(* Logix 5000 project; controller MV vendor 1 type 14 code 217 rev 31.11; software revision 31.00; part 2 of 53 *)

   MC_N224 : INT[255] := ([0] := 70, [1] := 59, [2] := 96, [3] := -32768, [4] := 9999, [5] := 9999, [6] := 9999, [7] := -32768);   // P24 CHECK CIP program 24 plant item check list
   MC_N225 : INT[255] := ([0] := 70, [1] := 59, [2] := 96, [3] := -32768, [4] := 9999, [5] := 9999, [6] := 9999, [7] := -32768);   // P25 CHECK CIP program 25 plant item check list
   MC_N226 : INT[255] := ([0] := 79, [1] := -32768, [2] := 9999, [3] := 9999, [4] := 9999, [5] := 9999, [6] := 9999, [7] := -32768);   // P26 CHECK CIP program 26 plant item check list
   MC_N227 : INT[255] := ([0] := 62, [1] := 99, [2] := -32768, [3] := 9999, [4] := 9999, [5] := 9999, [6] := 9999, [7] := -32768);   // P27 CHECK CIP program 27 plant item check list
   MC_N228 : INT[255] := ([0] := 61, [1] := 98, [2] := -32768, [3] := 9999, [4] := 9999, [5] := 9999, [6] := 9999, [7] := -32768);   // P28 CHECK CIP program 28 plant item check list
   MC_N229 : INT[255] := ([0] := 60, [1] := 97, [2] := -32768, [3] := 9999, [4] := 9999, [5] := 9999, [6] := 9999, [7] := -32768);   // P29 CHECK CIP program 29 plant item check list
   MC_N23 : INT[255] := ([0] := -31733, [2] := 1500, [3] := 5, [7] := 5000, [11] := 100, [12] := 10, [13] := 20, [14] := 7, [15] := 1493, [17] := -819, [18] := 25828, [21] := 5042, [22] := 1500, [24] := 1500, [25] := 13106, [27] := 1500, [31] := 3, [34] := 23, [36] := 1493);   // P2 FLOW Control block and da ta for P2 flowrate P ID loop
        [37]   // P2 flowrate PID saved op.mode
        [31].1   // P2 flowrate PID loop high absolute alarm flag
        [14]   // P2 flowrate PID loop process variable
        [31].0   // P2 flowrate PID loop deviation alarm flag
        [28]   // P2 flowrate PID loop high absolute alarm setting
        [31].2   // P2 flowrate PID loop low absolute alarm flag
        [30]   // P2 flowrate PID loop deviation alarm setting
        [38]   // P2 flowrate PID saved PLC output
        [26]   // P2 flowrate PID loop PLC output
        [25]   // P2 flowrate PID loop local (PC) output
        [0].1   // P2 flowrate PID loop auto/manual flag
        [2]   // P2 flowrate PID loop setpoint
        [27]   // P2 flowrate PID loop PLC setpoint
        [29]   // P2 flowrate PID loop low absolute alarm setting
        [35]   // P2 flowrate PID loop desired output
        [23]   // P2 flow op.mode: 0: PLC manual; 1: PLC setpoint; 2: Local manual; 3: Local setpoint;
        [36]   // Work register
   MC_N230 : INT[255] := ([0] := 60, [1] := 97, [2] := -32768, [3] := 9999, [4] := 9999, [5] := 9999, [6] := 9999, [7] := -32768);   // P30 CHECK CIP program 30 plant item check list
   MC_N231 : INT[255] := ([0] := 60, [1] := 97, [2] := -32768, [3] := 9999, [4] := 9999, [5] := 9999, [6] := 9999, [7] := -32768);   // P31 CHECK CIP program 31 plant item check list
   MC_N232 : INT[255] := ([0] := 60, [1] := 97, [2] := -32768, [3] := 9999, [4] := 9999, [5] := 9999, [6] := 9999, [7] := -32768);   // P32 CHECK CIP program 32 plant item check list
   MC_N233 : INT[255] := ([0] := 59, [1] := 96, [2] := -32768, [3] := 9999, [4] := 9999, [5] := 9999, [6] := 9999, [7] := -32768);   // P33 CHECK CIP program 33 plant item check list
   MC_N234 : INT[255] := ([0] := 59, [1] := 96, [2] := -32768, [3] := 9999, [4] := 9999, [5] := 9999, [6] := 9999, [7] := -32768);   // P34 CHECK CIP program 34 plant item check list
   MC_N235 : INT[255] := ([0] := 59, [1] := 96, [2] := -32768, [3] := 9999, [4] := 9999, [5] := 9999, [6] := 9999, [7] := -32768);   // P35 CHECK CIP program 35 plant item check list
   MC_N236 : INT[255] := ([0] := 59, [1] := 96, [2] := -32768, [3] := 9999, [4] := 9999, [5] := 9999, [6] := 9999, [7] := -32768);   // P36 CHECK CIP program 36 plant item check list
   MC_N237 : INT[255] := ([0] := 59, [1] := 96, [2] := -32768, [3] := 9999, [4] := 9999, [5] := 9999, [6] := 9999, [7] := -32768);   // P37 CHECK CIP program 37 plant item check list
   MC_N238 : INT[255] := ([0] := 59, [1] := 96, [2] := -32768, [3] := 9999, [4] := 9999, [5] := 9999, [6] := 9999, [7] := -32768);   // P38 CHECK CIP program 38 plant item check list
   MC_N239 : INT[255] := ([0] := 59, [1] := 96, [2] := -32768, [3] := 9999, [4] := 9999, [5] := 9999, [6] := 9999, [7] := -32768);   // P39 CHECK CIP program 39 plant item check list
   MC_N245 : INT[255];   // CC_WORK Continuous checking program work area
        [4].11   // CW deenergised input flag
        [6]   // Checking timer accumulator mask
        [15].0   // Current checkword is unused flag
        [2]   // Current item's energised input pointer
        [1]   // Current item's output pointer
        [3]   // Current item's Deenergised input pointer
        [4].10   // CW energised input flag
        [10].0   // Checking scan enabled flag
        [4].9   // CW desired output flag
        [0]   // Checkword pointer
        [16]   // Output slot update counter
        [28]   // No.items checked this scan
        [4]   // Current item's checkword
        [4].13   // CW checking inhibit flag
        [27]   // No new faults counter
        [4].12   // CW cycle flag
        [4].15   // CW fault flag
        [4].8   // CW manual flag
   MC_N255 : INT[255] := ([0] := 2208, [1] := 2208, [2] := 2208, [3] := 2208, [4] := 2208, [5] := 1696, [6] := 2208, [7] := 2208, [8] := 2208, [9] := 2208, [10] := 2208, [11] := 1696, [12] := 2208, [13] := 2208, [14] := 1696, [15] := 2112, [16] := 1600, [17] := 2112, [18] := 2112, [19] := 10304, [20] := 2112, [21] := 2112, [22] := 2112, [23] := 2112, [24] := 2112, [25] := 10304, [26] := 2112, [27] := 2112, [28] := 2112, [29] := 2112, [30] := 2112, [31] := 2112, [32] := 2112, [33] := 2112, [34] := 2112, [35] := 2112, [36] := 2112, [37] := 2112, [38] := 2112, [39] := 2112, [40] := 2112, [41] := 2112, [42] := 2112, [43] := 2112, [44] := 2112, [45] := 2112, [46] := 2112, [47] := 2112, [48] := 2112, [49] := 2112, [50] := 2112, [51] := 2112, [52] := 8256, [53] := 8256, [55] := 8256, [56] := 2112, [59] := 2112, [60] := 2112, [61] := 2112, [62] := 2112,
        [63] := 2112, [64] := 1600, [65] := 2112, [66] := 1600, [67] := 2112, [68] := 2112, [69] := 2112, [70] := 2112, [71] := 2112, [72] := 2112, [73] := 2112, [74] := 2112, [75] := 2112, [76] := 2112, [77] := 2112, [78] := 2112, [79] := 2112, [96] := 1600, [97] := 1600, [98] := 1600, [99] := 1600);   // CHECKWORDS Plant item checkword s
   MC_N7 : INT[255] := ([0] := 23, [1] := 22, [2] := 28, [4] := 2005, [5] := 5, [6] := 563, [7] := 84, [8] := 657, [9] := 653, [10] := -1);   // INTEGER
        [6]   // CH1/PTX scaled input
        [7]   // CH2/PTX scaled input
        [2]   // CH1/CTX1 scaled input
        [3]   // CH2/CTX2 scaled input
        [0]   // DT1 CTX-001 scaled input
        [1]   // DT2 CTX-002 scaled input
        [8]   // DT1 TTX-001 scaled input
        [9]   // DT2 TTX-002 scaled input
        [10]   // CH2/FM FV Bypass scaled input
        [4]   // CH1/FM scaled input
        [5]   // CH2/FM scaled input
   MC_N80 : INT[255] := ([0] := 5, [1] := 50, [2] := 4, [6] := 3, [7] := 23, [8] := 650, [10] := -1, [11] := 1, [13] := 10800, [14] := 1, [17] := 50, [18] := 7, [19] := 1, [20] := 2, [21] := 18);   // SRV1_PLC Detergent tank 1 ser vice PLC data
        [13]   // SV1 event register
        [21].1   // Channel 1 DT1 in use flag
        [21].3   // Channel 2 DT1 in use flag
        [2].0   // DT1 service manual start button available
        [2].15   // DT1 service command update toggle flag
        [21].4   // CH1/DT1 maintain temp.during service flag
        [21].5   // CH2/DT1 maintain temp.during service flag
        [20]   // DT1 service command processor current step
        [2].4   // DT1 service abort button available
        [21].0   // CH1 request DT1 service flag
        [21].2   // CH2 request DT1 service flag
        [8]   // DT1 service target detergent temp.
        [2].1   // DT1 manual service startup in progress
        [18].8   // DT1 service drive caustic pump flag
        [18].0   // DT1 service active flag
        [32].0   // DT1 service start by boilerhouse OSR
        [2].3   // DT1 service continue button available
        [6].0   // DT1 detergent strength ok
        [10]   // DT1 service routine fault register
        [18].1   // DT1 automatic service flag
        [6].1   // DT1 detergent temperature ok
        [17]   // DT1 service restart step
        [18].2   // DT1 service complete
        [6].2   // DT1 detergent diluted
        [11]   // SV1 fault parameter #1
        [12]   // SV1 fault parameter #2
        [14]   // SV1 event parameter #1
        [15]   // SV1 event parameter #2
        [1]   // DT1 service current step
        [2].2   // DT1 service stop button available
        [7]   // DT1 service target detergent strength
        [18].14   // Reset DT1 service flag
        [0]   // DT1 Service status 0:Unavailable; 1:Idle; 2:Running; 3:Stopped; 4:Faulted 5: Automatic
   MC_N80_10_alarm : ALARM_DIGITAL;
   MC_N80_10_Alarm_Ready : BOOL;
   MC_N80_10_Delayed_Timer2 : TIMER := (PRE := 1000);
   MC_N80_10_Fault_Returned : STRING;
   MC_N80_10_SQL_Done : DINT := -1;
   MC_N80_13_alarm : ALARM_DIGITAL;
   MC_N80_13_Alarm_Ready : BOOL := 1;
   MC_N80_13_Delayed_Timer2 : TIMER := (PRE := 1000);
   MC_N80_13_Event_Returned : STRING := 'Detergent tank service complete.';
   MC_N80_13_SQL_Done : DINT := -1;
   MC_N80_19_0_Storagebit : BOOL;
   MC_N81 : INT[255];   // SV1_PC Detergent tank 1 ser vice PC to PLC data
        [0].2   // Stop DT1 service
        [0].15   // DT1 manual service startup cancelled
        [0].0   // DT1 initiate manual service startup
        [0].4   // Abort DT1 service
        [0].1   // Start DT1 manual service
        [0]   // DT1 service PC button selected
        [0].3   // Continue DT1 service
   MC_N82 : INT[255] := ([0] := 14, [1] := 16, [2] := 34, [3] := 36, [4] := 41, [5] := 43, [6] := 45, [7] := 66, [8] := 78, [9] := -32768, [10] := 9999, [11] := 9999, [12] := 9999, [13] := 9999, [14] := 9999, [15] := 9999);   // SV1 ITEMS Chwd.nos.of items to be checked for DT1 service
        [6]   // SV1 checkword no.
        [8]   // CP1 checkword no.
        [0]   // CH1/DR1 checkword no.
        [1]   // CH1/DT1 checkword no.
        [2]   // CH2/DR1 checkword no.
        [3]   // CH2/DT1 checkword no.
        [4]   // FL/D1 checkword no.
        [5]   // CD/T1 checkword no.
        [7]   // P3 checkword no.
   MC_N90 : INT[255] := ([0] := 1, [2] := -32767, [10] := -1, [11] := 2, [13] := 10800, [14] := 2);   // SV2_PLC Detergent tank 2 ser vice PLC data
        [13]   // SV2 event register
        [21].1   // Channel 1 DT2 in use flag
        [21].3   // Channel 2 DT2 in use flag
        [2].0   // DT2 service manual start button available
        [2].15   // DT2 service command update toggle flag
        [21].4   // CH1/DT2 maintain temp.during service flag
        [21].0   // CH1 request DT2 service flag
        [21].5   // CH2/DT2 maintain temp.during service flag
        [20]   // DT2 service command processor current step
        [21].2   // CH2 request DT2 service flag
        [8]   // DT2 service target detergent temp.
        [2].4   // DT2 service abort button available
        [18].0   // DT2 service active flag
        [2].1   // DT2 manual service startup in progress
        [32].0   // DT2 service start by boilerhouse OSR
        [18].8   // DT2 service drive caustic pump flag
        [2].3   // DT2 service continue button available
        [6].0   // DT2 detergent strength ok
        [10]   // DT2 service routine fault register
        [18].1   // DT2 automatic service flag
        [6].1   // DT2 detergent temperature ok
        [17]   // DT2 service restart step
        [18].2   // DT2 service complete
        [6].2   // DT2 detergent diluted
        [11]   // SV2 fault parameter #1
        [14]   // SV2 event parameter #1
        [1]   // DT2 service current step
        [2].2   // DT2 service stop button available
        [7]   // DT2 service target detergent strength
        [18].14   // Reset DT2 service flag
        [0]   // DT2 Service status 0:Unavailable; 1:Idle; 2:Running; 3:Stopped; 4:Faulted 5: Automatic
   MC_N90_10_alarm : ALARM_DIGITAL;
   MC_N90_10_Alarm_Ready : BOOL;
   MC_N90_10_Delayed_Timer2 : TIMER := (PRE := 1000);
   MC_N90_10_Fault_Returned : STRING;
   MC_N90_10_SQL_Done : DINT := -1;
   MC_N90_13_alarm : ALARM_DIGITAL;
   MC_N90_13_Alarm_Ready : BOOL := 1;
   MC_N90_13_Delayed_Timer2 : TIMER := (PRE := 1002);
   MC_N90_13_Event_Returned : STRING := 'Detergent tank service complete.';
   MC_N90_13_SQL_Done : DINT := -1;
   MC_N90_19_0_Storagebit : BOOL;
   MC_N90_32_0_Storagebit : BOOL;
   MC_N91 : INT[255];   // SV2_PC Detergent tank 2 ser vice PC to PLC data
        [0].2   // Stop DT2 service
        [0].15   // DT2 manual service startup cancelled
        [0].0   // DT2 initiate manual service startup
        [0].4   // Abort DT2 service
        [0].1   // Start DT2 manual service
        [0]   // DT2 service PC button selected
        [0].3   // Continue DT2 service
   MC_N92 : INT[255] := ([0] := 15, [1] := 17, [2] := 35, [3] := 37, [4] := 42, [5] := 44, [6] := 46, [7] := 67, [8] := 78, [9] := -32768, [10] := 9999, [11] := 9999, [12] := 9999, [13] := 9999, [14] := 9999, [15] := 9999);   // SV2 ITEMS Chwd.nos.of items to be checked for DT2 service
        [6]   // SV2 checkword no.
        [8]   // CP1 checkword no.
        [0]   // CH1/DR2 checkword no.
        [1]   // CH1/DT2 checkword no.
        [2]   // CH2/DR2 checkword no.
        [3]   // CH2/DT2 checkword no.
        [4]   // FL/D2 checkword no.
        [7]   // P4 checkword no.
        [5]   // CD/T2 checkword no.
   MC_ONE_SEC : ALIAS FOR MC_T4[0].DN;
   MC_P1 : PlantItem := (CW := 2#0000_0000_0000_0001_0000_1100_1000_1011, CheckTime := 8, CheckTimer := 8, DriveBits := 1);   // P1
   MC_P1_ALARM : ALARM_DIGITAL;
   MC_P1_D : ALIAS FOR RIO_Rack_2:10:O.Data.0;
   MC_P1_Flow_PID : PID := (CTL := -2139061120, EN := 1, PE := 1, INI := 1, DVNA := 1, PVHA := 1, SP := 200.0, KP := 0.5, KI := 50.0, MAXS := 500.0, SO := 72.11798, MAXO := 100.0, MINO := 10.0, UPD := 1.0, PV := 200.53125, ERR := -0.53125, OUT := 72.11798, MAXI := 500.0, TIE := 72.118, MAXCV := 100.0, MAXTIE := 100.0, DATA[0] := 72.171104, DATA[1] := -641.7, DATA[2] := 200.53125, DATA[3] := -0.53125, DATA[4] := 200.0, DATA[5] := 0.2, DATA[6] := 1.0, DATA[7] := 16.0, DATA[8] := 0.5, DATA[9] := 50.0, DATA[11] := 0.5, DATA[12] := 0.00016666666, DATA[15] := 1.0, DATA[16] := 1.0);
   MC_P1_Flow_PID_Output : REAL := 72.16245;
   MC_P1_FPID_RESTORE : ALIAS FOR MC_N100[29].4;
   MC_P1_FPID_SAVE : ALIAS FOR MC_N100[29].3;
   MC_P1_PPID_RESTORE : ALIAS FOR MC_N100[29].2;
   MC_P1_PPID_SAVE : ALIAS FOR MC_N100[29].1;
   MC_P1_Pressure_PID : PID := (CTL := -2071952768, EN := 1, SWM := 1, PE := 1, INI := 1, DVPA := 1, PVHA := 1, SP := 65.0, KP := 1.0, KI := 2.0, MAXS := 150.0, MAXO := 100.0, UPD := 1.0, PV := 52.26563, ERR := 12.734371, MAXI := 150.0, MAXCV := 100.0, MAXTIE := 100.0, DATA[0] := -8.489581, DATA[1] := -557.50006, DATA[2] := 52.26563, DATA[3] := 12.734371, DATA[4] := 65.0, DATA[5] := 0.6666667, DATA[6] := 1.0, DATA[7] := 16.0, DATA[8] := 1.0, DATA[9] := 2.0, DATA[11] := 1.0, DATA[12] := 0.008333334, DATA[15] := 1.0, DATA[16] := 1.0);
   MC_P1_Pressure_PID_Output : REAL;
   MC_P1_R : ALIAS FOR RIO_Rack_2:11:I.Data.0;
   MC_P1_SP_AO : PlantItem := (Scaled := 72.161766);   // P1_SP
   MC_P1_SP_AO_RawOutput : ALIAS FOR RIO_Rack_2:3:O.Ch0Data;   // Real Analog Input , Do Not Use In Code
   MC_P1_T : ALIAS FOR RIO_Rack_2:11:I.Data.15;
   MC_P2 : PlantItem := (CW := 2#0000_0000_0000_0000_0000_1100_0000_0000, CheckTime := 8, CheckTimer := 8);   // P2
   MC_P2_ALARM : ALARM_DIGITAL;
   MC_P2_D : ALIAS FOR RIO_Rack_2:10:O.Data.1;
   MC_P2_Flow_PID : PID := (CTL := -2071952768, EN := 1, SWM := 1, PE := 1, INI := 1, DVPA := 1, PVHA := 1, SP := 150.0, KP := 0.5, KI := 50.0, MAXS := 500.0, MAXO := 100.0, UPD := 1.0, PV := 1.0, ERR := 149.0, MAXI := 500.0, MAXCV := 100.0, MAXTIE := 100.0, DATA[0] := -14.900001, DATA[1] := -3.2, DATA[2] := 1.0, DATA[3] := 149.0, DATA[4] := 150.0, DATA[5] := 0.2, DATA[6] := 1.0, DATA[7] := 16.0, DATA[8] := 0.5, DATA[9] := 50.0, DATA[11] := 0.5, DATA[12] := 0.00016666666, DATA[15] := 1.0, DATA[16] := 1.0);
   MC_P2_Flow_PID_Output : REAL;
   MC_P2_FPID_RESTORE : ALIAS FOR MC_N120[29].4;
   MC_P2_FPID_SAVE : ALIAS FOR MC_N120[29].3;
   MC_P2_PPID_RESTORE : ALIAS FOR MC_N120[29].2;
   MC_P2_PPID_SAVE : ALIAS FOR MC_N120[29].1;
   MC_P2_Pressure_PID : PID := (CTL := -2071952768, EN := 1, SWM := 1, PE := 1, INI := 1, DVPA := 1, PVHA := 1, SP := 45.0, KP := 0.1, KI := 2.0, MAXS := 150.0, MAXO := 100.0, UPD := 1.0, PV := 8.3625, ERR := 36.6375, MAXI := 150.0, MAXCV := 100.0, MAXTIE := 100.0, DATA[0] := -2.4425, DATA[1] := -89.200005, DATA[2] := 8.3625, DATA[3] := 36.6375, DATA[4] := 45.0, DATA[5] := 0.6666667, DATA[6] := 1.0, DATA[7] := 16.0, DATA[8] := 0.1, DATA[9] := 2.0, DATA[11] := 0.1, DATA[12] := 0.00083333335, DATA[15] := 1.0, DATA[16] := 1.0);
   MC_P2_Pressure_PID_Output : REAL;
   MC_P2_R : ALIAS FOR RIO_Rack_2:11:I.Data.1;
   MC_P2_SP_AO : PlantItem;   // P2_SP
   MC_P2_SP_AO_RawOutput : ALIAS FOR RIO_Rack_2:3:O.Ch1Data;   // Real Analog Input , Do Not Use In Code
   MC_P2_T : ALIAS FOR RIO_Rack_2:11:I.Data.16;
   MC_P3 : PlantItem := (CW := 2#0000_0000_0000_0000_0000_1100_1000_1011, CheckTime := 8, CheckTimer := 8, DriveBits := 1);   // P3
   MC_P3_ALARM : ALARM_DIGITAL;
   MC_P3_D : ALIAS FOR RIO_Rack_2:10:O.Data.2;
   MC_P3_R : ALIAS FOR RIO_Rack_2:11:I.Data.2;
   MC_P4 : PlantItem := (CW := 2#0000_0000_0000_0000_0000_1100_0000_0000, CheckTime := 8, CheckTimer := 8);   // P4
   MC_P4_ALARM : ALARM_DIGITAL;
   MC_P4_D : ALIAS FOR RIO_Rack_2:10:O.Data.3;
   MC_P4_R : ALIAS FOR RIO_Rack_2:11:I.Data.3;
   MC_PILZ : PlantItem := (CW := 2#0000_0000_0000_0100_0000_0000_0000_0001);   // PILZ
   MC_PILZ_RawInput : ALIAS FOR RIO_Rack_2:12:I.Data.31;   // MC_PILZ
   MC_PROXY2 : PlantItem;   // PROXY2
   MC_PROXY2_RawInput : ALIAS FOR RIO_Rack_2:12:I.Data.30;   // MC_PROXY2
   MC_PROXY_RawInput : ALIAS FOR RIO_Rack_2:12:I.Data.14;   // MC_PROXY
   MC_PX_100 : PlantItem;   // PX_100
   MC_PX_100_RawInput : ALIAS FOR RIO_Rack_2:11:I.Data.18;   // MC_PX_100
   MC_PX_101 : PlantItem;   // PX_101
   MC_PX_101_RawInput : ALIAS FOR RIO_Rack_2:11:I.Data.19;   // MC_PX_101
   MC_R2_SW1 : PlantItem;   // R2_SW1
   MC_R2_SW1_RawInput : ALIAS FOR RIO_Rack_2:12:I.Data.0;   // MC_R2_SW1
   MC_R2_SW2 : PlantItem;   // R2_SW2
   MC_R2_SW2_RawInput : ALIAS FOR RIO_Rack_2:12:I.Data.1;   // MC_R2_SW2
   MC_R2_SW3 : PlantItem;   // R2_SW3
   MC_R2_SW3_1 : PlantItem;   // R2_SW3_1
   MC_R2_SW3_1_RawInput : ALIAS FOR RIO_Rack_2:12:I.Data.3;   // MC_R2_SW3_1
   MC_R2_SW3_RawInput : ALIAS FOR RIO_Rack_2:12:I.Data.2;   // MC_R2_SW3
   MC_R2_SW4 : PlantItem := (CW := 2#0000_0000_0000_0100_0000_0000_0000_0001);   // R2_SW4
   MC_R2_SW4_RawInput : ALIAS FOR RIO_Rack_2:12:I.Data.4;   // MC_R2_SW4
   MC_R3_SW1 : PlantItem;   // R3_SW1
   MC_R3_SW1_RawInput : ALIAS FOR RIO_Rack_2:12:I.Data.5;   // MC_R3_SW1
   MC_R3_SW2 : PlantItem;   // R3_SW2
   MC_R3_SW2_1 : PlantItem := (CW := 2#0000_0000_0000_0100_0000_0000_0010_0001);   // PROXY
   MC_R3_SW2_RawInput : ALIAS FOR RIO_Rack_2:12:I.Data.6;   // MC_R3_SW2
   MC_R3_SW3 : PlantItem;   // R3_SW3
   MC_R3_SW3_1 : ALIAS FOR MC_N112[9].1;
   MC_R3_SW3_2 : ALIAS FOR MC_N112[9].0;
   MC_R3_SW3_3 : ALIAS FOR MC_N112[9].2;
   MC_R3_SW3_RawInput : ALIAS FOR RIO_Rack_2:12:I.Data.7;   // MC_R3_SW3
   MC_R3R_C_ALARM : ALARM_DIGITAL;
   MC_R3R_DR : PlantItem := (CW := 2#0000_0000_0000_0000_0000_0000_0001_0000, CheckTime := 8, CheckTimer := 15);   // R3R_DR
   MC_R3R_DR_ALARM : ALARM_DIGITAL;
   MC_R3R_DR_C : ALIAS FOR RIO_Rack_2:9:I.Data.20;
   MC_R3R_DR_DR : ALIAS FOR RIO_Rack_2:8:O.Data.24;
   MC_R3R_DR_O : ALIAS FOR RIO_Rack_2:9:I.Data.16;
   MC_R3R_O_ALARM : ALARM_DIGITAL;
   MC_R3S_C_ALARM : ALARM_DIGITAL;
   MC_R3S_DR : PlantItem := (CW := 2#0000_0000_0000_0000_0000_0001_0000_0000, CheckTime := 8, CheckTimer := 15);   // R3S_DR
   MC_R3S_DR_ALARM : ALARM_DIGITAL;
   MC_R3S_DR_C : ALIAS FOR RIO_Rack_2:9:I.Data.15;
   MC_R3S_DR_DR : ALIAS FOR RIO_Rack_2:8:O.Data.23;
   MC_R3S_DR_O : ALIAS FOR RIO_Rack_2:9:I.Data.11;
   MC_R3S_O_ALARM : ALARM_DIGITAL;
   MC_R3V1 : PlantItem := (CW := 2#0000_0000_0000_0000_0000_0001_0000_0000, CheckTime := 8, CheckTimer := 15);   // R3V1
   MC_R3V1_ALARM : ALARM_DIGITAL;
   MC_R3V1_C : ALIAS FOR RIO_Rack_2:9:I.Data.12;
   MC_R3V1_DR : ALIAS FOR RIO_Rack_2:8:O.Data.20;
   MC_R3V1_O : ALIAS FOR RIO_Rack_2:9:I.Data.8;
   MC_R3V2 : PlantItem := (CW := 2#0000_0000_0000_0000_0000_0001_0000_0000, CheckTime := 8, CheckTimer := 15);   // R3V2
   MC_R3V2_ALARM : ALARM_DIGITAL;
   MC_R3V2_C : ALIAS FOR RIO_Rack_2:9:I.Data.13;
   MC_R3V2_DR : ALIAS FOR RIO_Rack_2:8:O.Data.21;
   MC_R3V2_O : ALIAS FOR RIO_Rack_2:9:I.Data.9;
   MC_R3V3_C : ALIAS FOR RIO_Rack_2:9:I.Data.14;
   MC_R3V3_O : ALIAS FOR RIO_Rack_2:9:I.Data.10;
   MC_R4_SW1 : PlantItem;   // R4_SW1
   MC_R4_SW1_RawInput : ALIAS FOR RIO_Rack_2:12:I.Data.8;   // MC_R4_SW1
   MC_R4_SW2 : PlantItem;   // R4_SW2
   MC_R4_SW2_RawInput : ALIAS FOR RIO_Rack_2:12:I.Data.9;   // MC_R4_SW2
   MC_R4_SW3 : PlantItem := (CW := 2#0000_0000_0000_0100_0000_0000_0000_0001);   // R4_SW3
   MC_R4_SW3_RawInput : ALIAS FOR RIO_Rack_2:12:I.Data.10;   // MC_R4_SW3
   MC_R4_SW4 : PlantItem;   // R4_SW4
   MC_R4_SW4_RawInput : ALIAS FOR RIO_Rack_2:12:I.Data.11;   // MC_R4_SW4
   MC_R4_SW6 : PlantItem := (CW := 2#0000_0000_0000_0100_0000_0000_0000_0001);   // R4_SW6
   MC_R4_SW6_RawInput : ALIAS FOR RIO_Rack_2:12:I.Data.12;   // MC_R4_SW6
   MC_R6_SW1 : PlantItem := (CW := 2#0000_0000_0000_0100_0000_0000_0000_0001);   // R6_SW1
   MC_R6_SW1_RawInput : ALIAS FOR RIO_Rack_2:12:I.Data.13;   // MC_R6_SW1
   MC_RackingTanks_Emptying_event : STRING;
   MC_RackingTanks_Emptying_event_prefix : STRING;
   MC_RackingTanks_Filling_event : STRING;
   MC_RackingTanks_Filling_event_prefix : STRING;
   MC_RT_Emptying_Log_ID : DINT := 1;
   MC_RT_Filling_Log_ID : DINT := 2;
   MC_SFile : INT[255] := ([4] := -19490, [37] := 2020, [40] := 17, [42] := 5);   // SLC Equivalent System File, So Original Code Can Remain
        [40]   // Clock Calendar Hours
        [1].15   // First Scan Flag
        [41]   // Clock Calendar Minutes
   MC_SP_R1_1 : PlantItem := (CW := 2#0000_0000_0000_0000_0000_1100_0000_0000, CheckTime := 8, CheckTimer := 8);   // SP_R1_1
   MC_SP_R1_1_ALARM : ALARM_DIGITAL;
   MC_SP_R1_1_D : ALIAS FOR RIO_Rack_2:10:O.Data.4;
   MC_SP_R1_1_R : ALIAS FOR RIO_Rack_2:11:I.Data.4;
   MC_SP_R2_1 : PlantItem := (CW := 2#0000_0000_0000_0000_0000_1100_0000_0000, CheckTime := 8, CheckTimer := 8);   // SP_R2_1
   MC_SP_R2_1_ALARM : ALARM_DIGITAL;
   MC_SP_R2_1_D : ALIAS FOR RIO_Rack_2:10:O.Data.5;
   MC_SP_R2_1_R : ALIAS FOR RIO_Rack_2:11:I.Data.5;
   MC_SP_R2_2 : PlantItem := (CW := 2#0000_0000_0000_0000_0000_1100_0000_0000, CheckTime := 8, CheckTimer := 8);   // SP_R2_2
   MC_SP_R2_2_ALARM : ALARM_DIGITAL;
   MC_SP_R2_2_D : ALIAS FOR RIO_Rack_2:10:O.Data.15;
   MC_SP_R2_2_R : ALIAS FOR RIO_Rack_2:11:I.Data.14;
   MC_SP_R3_1 : PlantItem := (CW := 2#0000_0000_0000_0000_0000_1100_0000_0000, CheckTime := 8, CheckTimer := 8);   // SP_R3_1
   MC_SP_R3_1_ALARM : ALARM_DIGITAL;
   MC_SP_R3_1_D : ALIAS FOR RIO_Rack_2:10:O.Data.6;
   MC_SP_R3_1_R : ALIAS FOR RIO_Rack_2:11:I.Data.6;
   MC_SP_R5_1 : PlantItem := (CW := 2#0000_0000_0000_0000_0000_1100_0000_0000, CheckTime := 8, CheckTimer := 8);   // SP_R5_1
   MC_SP_R5_1_ALARM : ALARM_DIGITAL;
   MC_SP_R5_1_D : ALIAS FOR RIO_Rack_2:10:O.Data.7;
   MC_SP_R5_1_R : ALIAS FOR RIO_Rack_2:11:I.Data.7;
   MC_SP_R5_2 : PlantItem := (CW := 2#0000_0000_0000_0000_0000_1100_0000_0000, CheckTime := 8, CheckTimer := 8);   // SP_R5_2
   MC_SP_R5_2_ALARM : ALARM_DIGITAL;
   MC_SP_R5_2_D : ALIAS FOR RIO_Rack_2:10:O.Data.8;
   MC_SP_R5_2_R : ALIAS FOR RIO_Rack_2:11:I.Data.8;
   MC_SP_R6_1 : PlantItem := (CW := 2#0000_0000_0000_0000_0000_1100_0000_0000, CheckTime := 8, CheckTimer := 8);   // SP_R6_1
   MC_SP_R6_1_ALARM : ALARM_DIGITAL;
   MC_SP_R6_1_D : ALIAS FOR RIO_Rack_2:10:O.Data.9;
   MC_SP_R6_1_R : ALIAS FOR RIO_Rack_2:11:I.Data.9;
   MC_SP_R6_2 : PlantItem := (CW := 2#0000_0000_0000_0000_0000_1100_0000_0000, CheckTime := 8, CheckTimer := 8);   // SP_R6_2
   MC_SP_R6_2_ALARM : ALARM_DIGITAL;
   MC_SP_R6_2_D : ALIAS FOR RIO_Rack_2:10:O.Data.10;
   MC_SP_R6_2_R : ALIAS FOR RIO_Rack_2:11:I.Data.10;
   MC_SP_R6_3 : PlantItem := (CW := 2#0000_0000_0000_0000_0000_1100_0000_0000, CheckTime := 8, CheckTimer := 8);   // SP_R6_3
   MC_SP_R6_3_ALARM : ALARM_DIGITAL;
   MC_SP_R6_3_D : ALIAS FOR RIO_Rack_2:10:O.Data.11;
   MC_SP_R6_3_R : ALIAS FOR RIO_Rack_2:11:I.Data.11;
   MC_SP_R6_4 : PlantItem := (CW := 2#0000_0000_0000_0000_0000_1100_0000_0000, CheckTime := 8, CheckTimer := 8);   // SP_R6_4
   MC_SP_R6_4_ALARM : ALARM_DIGITAL;
   MC_SP_R6_4_D : ALIAS FOR RIO_Rack_2:10:O.Data.12;
   MC_SP_R6_4_R : ALIAS FOR RIO_Rack_2:11:I.Data.12;
   MC_SP_R6_5 : PlantItem := (CW := 2#0000_0000_0000_0000_0000_1100_0000_0000, CheckTime := 8, CheckTimer := 8);   // SP_R6_5
   MC_SP_R6_5_ALARM : ALARM_DIGITAL;
   MC_SP_R6_5_D : ALIAS FOR RIO_Rack_2:10:O.Data.13;
   MC_SP_R6_5_R : ALIAS FOR RIO_Rack_2:11:I.Data.13;
   MC_SP_V12TO17 : PlantItem;   // SP_V12TO17
   MC_SP_V12TO17_RawOutput : ALIAS FOR RIO_Rack_2:10:O.Data.17;   // MC_SP_V12TO17
   MC_SPV1 : PlantItem := (CW := 2#0000_0000_0000_0000_0000_0000_0001_0000, CheckTime := 8, CheckTimer := 8);   // SPV1
   MC_SPV1_ALARM : ALARM_DIGITAL;
   MC_SPV1_C : ALIAS FOR RIO_Rack_2:7:I.Data.31;
   MC_SPV1_DR : ALIAS FOR RIO_Rack_2:8:O.Data.15;
   MC_SPV1_O : ALIAS FOR RIO_Rack_2:7:I.Data.27;
   MC_SPV2 : PlantItem := (CW := 2#0000_0000_0000_0000_0000_0000_0001_0000, CheckTime := 8, CheckTimer := 8);   // SPV2
   MC_SPV2_ALARM : ALARM_DIGITAL;
   MC_SPV2_C : ALIAS FOR RIO_Rack_2:9:I.Data.4;
   MC_SPV2_DR : ALIAS FOR RIO_Rack_2:8:O.Data.16;
   MC_SPV2_O : ALIAS FOR RIO_Rack_2:9:I.Data.0;
   MC_SPV3 : PlantItem := (CW := 2#0000_0000_0000_0000_0000_0000_0001_0000, CheckTime := 8, CheckTimer := 8);   // SPV3
   MC_SPV3_ALARM : ALARM_DIGITAL;
   MC_SPV3_C : ALIAS FOR RIO_Rack_2:9:I.Data.5;
   MC_SPV3_DR : ALIAS FOR RIO_Rack_2:8:O.Data.17;
   MC_SPV3_O : ALIAS FOR RIO_Rack_2:9:I.Data.1;
   MC_SPV4 : PlantItem := (CW := 2#0000_0000_0000_0000_0000_0000_0001_0000, CheckTime := 8, CheckTimer := 8);   // SPV4
   MC_SPV4_ALARM : ALARM_DIGITAL;
   MC_SPV4_C : ALIAS FOR RIO_Rack_2:9:I.Data.6;
   MC_SPV4_DR : ALIAS FOR RIO_Rack_2:8:O.Data.18;
   MC_SPV4_O : ALIAS FOR RIO_Rack_2:9:I.Data.2;
   MC_SPV5 : PlantItem := (CW := 2#0000_0000_0000_0000_0000_0000_0001_0000, CheckTime := 8, CheckTimer := 8);   // SPV5
   MC_SPV5_ALARM : ALARM_DIGITAL;
   MC_SPV5_C : ALIAS FOR RIO_Rack_2:9:I.Data.7;
   MC_SPV5_DR : ALIAS FOR RIO_Rack_2:8:O.Data.19;
   MC_SPV5_O : ALIAS FOR RIO_Rack_2:9:I.Data.3;
   MC_SRV1_Log_ID : DINT := 54;
   MC_SRV2_Log_ID : DINT := 55;
   MC_SV1 : PlantItem := (CW := 2#0000_0000_0000_0000_0000_0000_0001_0000, CheckTime := 8, CheckTimer := 8);   // SV1
   MC_SV1_ACTIVE : ALIAS FOR MC_N80[18].0;   // DT1 service active flag
   MC_SV1_ALARM : ALARM_DIGITAL;
   MC_SV1_AUTO : ALIAS FOR MC_N80[18].1;   // DT1 automatic service flag
   MC_SV1_C : ALIAS FOR RIO_Rack_2:7:I.Data.29;
   MC_SV1_CSTEP : ALIAS FOR MC_N80[20];   // DT1 service command processor current step
   MC_SV1_DR : ALIAS FOR RIO_Rack_2:8:O.Data.13;
   MC_SV1_EVENT : ALIAS FOR MC_N80[13];   // SV1 event register
   MC_SV1_FAULT : ALIAS FOR MC_N80[10];   // DT1 service routine fault register
   MC_SV1_INIT : ALIAS FOR MC_N80[19].0;
   MC_SV1_O : ALIAS FOR RIO_Rack_2:7:I.Data.25;
   MC_SV1_RESET : ALIAS FOR MC_N80[18].14;   // Reset DT1 service flag
   MC_SV1_RESTART : ALIAS FOR MC_N80[17];   // DT1 service restart step
   MC_SV1_STATUS : ALIAS FOR MC_N80[0];   // DT1 Service status 0:Unavailable; 1:Idle; 2:Running; 3:Stopped; 4:Faulted 5: Automatic
   MC_SV1_STEP : ALIAS FOR MC_N80[1];   // DT1 service current step
   MC_SV2 : PlantItem := (CW := 2#0000_0000_0000_0000_0000_0000_0001_0000, CheckTime := 8, CheckTimer := 8);   // SV2
   MC_SV2_ACTIVE : ALIAS FOR MC_N90[18].0;   // DT2 service active flag
   MC_SV2_ALARM : ALARM_DIGITAL;
   MC_SV2_AUTO : ALIAS FOR MC_N90[18].1;   // DT2 automatic service flag
   MC_SV2_C : ALIAS FOR RIO_Rack_2:7:I.Data.30;
   MC_SV2_CSTEP : ALIAS FOR MC_N90[20];   // DT2 service command processor current step
   MC_SV2_DR : ALIAS FOR RIO_Rack_2:8:O.Data.14;
   MC_SV2_EVENT : ALIAS FOR MC_N90[13];   // SV2 event register
   MC_SV2_FAULT : ALIAS FOR MC_N90[10];   // DT2 service routine fault register
   MC_SV2_INIT : ALIAS FOR MC_N90[19].0;
   MC_SV2_O : ALIAS FOR RIO_Rack_2:7:I.Data.26;
   MC_SV2_RESET : ALIAS FOR MC_N90[18].14;   // Reset DT2 service flag
   MC_SV2_RESTART : ALIAS FOR MC_N90[17];   // DT2 service restart step
   MC_SV2_STATUS : ALIAS FOR MC_N90[0];   // DT2 Service status 0:Unavailable; 1:Idle; 2:Running; 3:Stopped; 4:Faulted 5: Automatic
   MC_SV2_STEP : ALIAS FOR MC_N90[1];   // DT2 service current step
   MC_T105 : TIMER[255] := ([0].PRE := 300000, [1].PRE := 10000, [2].PRE := 900000, [2].ACC := 814203, [2].EN := 1, [2].TT := 1, [5].PRE := 90000, [6].PRE := 120000, [7].PRE := 5000, [7].ACC := 5000, [7].EN := 1, [7].DN := 1, [8].PRE := 10000, [8].ACC := 10001, [8].EN := 1, [8].DN := 1, [9].PRE := 10000, [10].PRE := 10000, [10].ACC := 10001, [10].EN := 1, [10].DN := 1, [11].PRE := 10000, [12].PRE := 2000, [12].ACC := 216, [12].EN := 1, [12].TT := 1, [14].PRE := 5000, [15].PRE := 10000, [16].PRE := 5000, [17].PRE := 5000, [17].ACC := 5001, [17].EN := 1, [17].DN := 1, [18].PRE := 5000, [19].PRE := 5000);   // CH1 TIMERS Channel 1 timers
        [9]   // CH1 return flow off debounce timer
        [4]   // CH1 return pump off delay timer
        [2].DN   // CH1 current cycle complete
        [0].DN   // CH1 startup guard timer done
        [1].DN   // CH1 program validation timed-out
        [10]   // CH1 detergent return on debounce timer
        [16].TT   // CH1 prerinse supply close delay active
        [15]   // CH1 delay return flow check on restart timer
        [11]   // CH1 detergent return off debounce timer
        [16]   // CH1 prerinse supply close delay timer
        [8]   // CH1 return flow on debounce timer
        [14].TT   // CH1 return pump restart delay active
        [3].DN   // CH1 return pump on delay done
        [17]   // CH1 return to detergent tank timer
        [6]   // CH1 detergent return check timer
        [18]   // CH1 return to prerinse tank timer
        [1]   // CH1 program validation guard timer
        [19]   // CH1 return to drain timer
        [5]   // CH1 return flow check timer
        [12]   // CH1 item checking timer
        [3]   // CH1 return pump on delay timer
        [14]   // CH1 delay return pump restart timer
        [7]   // CH1 supply pump on delay timer
        [12].DN   // CH1 item checking timer done
        [4].DN   // CH1 return pump off delay done
        [0]   // CH1 startup guard timer
        [2]   // CH1 current cycle timer
   MC_T125 : TIMER[255] := ([0].PRE := 300000, [1].PRE := 10000, [2].PRE := 90000, [3].PRE := 60000, [4].PRE := 10000, [5].PRE := 120000, [6].PRE := 125000, [7].PRE := 5000, [8].PRE := 10000, [9].PRE := 20000, [10].PRE := 10000, [11].PRE := 10000, [12].PRE := 2000, [14].PRE := 5000, [15].PRE := 10000, [16].PRE := 5000, [17].PRE := 5000, [18].PRE := 5000, [19].PRE := 5000, [20].PRE := 5000, [20].ACC := 5001, [20].EN := 1, [20].DN := 1, [21].PRE := 5000, [22].PRE := 5000, [22].ACC := 5001, [22].EN := 1, [22].DN := 1, [23].PRE := 5000, [24].PRE := 30000, [25].PRE := 10000, [26].PRE := 30000);   // CH2 TIMERS Channel 2 timers
        [9]   // CH2 return flow off debounce timer
        [4]   // CH2 return pump off delay timer
        [2].DN   // CH2 current cycle complete
        [0].DN   // CH2 startup guard timer done
        [10]   // CH2 detergent return on debounce timer
        [1].DN   // CH2 program validation timed-out
        [16].TT   // CH2 prerinse supply close delay active
        [11]   // CH2 detergent return off debounce timer
        [15]   // CH2 delay return flow check on restart timer
        [8]   // CH2 return flow on debounce timer
        [16]   // CH2 prerinse supply close delay timer
        [14].TT   // CH2 return pump restart delay active
        [3].DN   // CH2 return pump on delay done
        [17]   // CH2 return to detergent tank timer
        [18]   // CH2 return to prerinse tank timer
        [6]   // CH2 detergent return check timer
        [1]   // CH2 program validation guard timer
        [19]   // CH2 return to drain timer
        [5]   // CH2 return flow check timer
        [12]   // CH2 item checking timer
        [14]   // CH2 delay return pump restart timer
        [3]   // CH2 return pump on delay timer
        [7]   // CH2 supply pump on delay timer
        [0]   // CH2 startup guard timer
        [12].DN   // CH2 item checking timer done
        [4].DN   // CH2 return pump off delay done
        [2]   // CH2 current cycle timer